(* Logix 5000 project; controller MV vendor 1 type 14 code 217 rev 31.11; software revision 31.00; part 29 of 53 *)
(* tags used below, declared in another part *)
   active : BOOL;
   Alarm_Reset : BOOL;
   CWD : CHECKWORD_FLAGS;
   Default_Check_Time : DINT;
   Item_Faults_Are_Latched : BOOL;
   Item_Simulation_Flag : BOOL;
   MC_CD_T2 : PlantItem;   // CD_T2
   MC_CH1_R1 : PlantItem;   // CH1_R1
   MC_CH1_R1_ALARM : ALARM_DIGITAL;
   MC_CH1_R1_C : ALIAS FOR RIO_Rack_2:4:I.Data.4;
   MC_CH1_R1_DR : ALIAS FOR RIO_Rack_2:5:O.Data.0;
   MC_CH1_R1_O : ALIAS FOR RIO_Rack_2:4:I.Data.0;
   MC_CH1_R1R : PlantItem;   // CH1_R1R
   MC_CH1_R1R_ALARM : ALARM_DIGITAL;
   MC_CH1_R1R_C : ALIAS FOR RIO_Rack_2:4:I.Data.14;
   MC_CH1_R1R_DR : ALIAS FOR RIO_Rack_2:5:O.Data.6;
   MC_CH1_R1R_O : ALIAS FOR RIO_Rack_2:4:I.Data.10;
   MC_CH1_R2 : PlantItem;   // CH1_R2
   MC_CH1_R2_ALARM : ALARM_DIGITAL;
   MC_CH1_R2_C : ALIAS FOR RIO_Rack_2:4:I.Data.5;
   MC_CH1_R2_DR : ALIAS FOR RIO_Rack_2:5:O.Data.1;
   MC_CH1_R2_O : ALIAS FOR RIO_Rack_2:4:I.Data.1;
   MC_CH1_R3 : PlantItem;   // CH1_R3
   MC_CH1_R3_ALARM : ALARM_DIGITAL;
   MC_CH1_R3_C : ALIAS FOR RIO_Rack_2:4:I.Data.6;
   MC_CH1_R3_DR : ALIAS FOR RIO_Rack_2:5:O.Data.2;
   MC_CH1_R3_O : ALIAS FOR RIO_Rack_2:4:I.Data.2;
   MC_CH1_R4 : PlantItem;   // CH1_R4
   MC_CH1_R4_ALARM : ALARM_DIGITAL;
   MC_CH1_R4_C : ALIAS FOR RIO_Rack_2:4:I.Data.7;
   MC_CH1_R4_DR : ALIAS FOR RIO_Rack_2:5:O.Data.3;
   MC_CH1_R4_O : ALIAS FOR RIO_Rack_2:4:I.Data.3;
   MC_CH1_R5 : PlantItem;   // CH1_R5
   MC_CH1_R5_ALARM : ALARM_DIGITAL;
   MC_CH1_R5_C : ALIAS FOR RIO_Rack_2:4:I.Data.12;
   MC_CH1_R5_DR : ALIAS FOR RIO_Rack_2:5:O.Data.4;
   MC_CH1_R5_O : ALIAS FOR RIO_Rack_2:4:I.Data.8;
   MC_CH1_R6 : PlantItem;   // CH1_R6
   MC_CH1_R6_ALARM : ALARM_DIGITAL;
   MC_CH1_R6_C : ALIAS FOR RIO_Rack_2:4:I.Data.13;
   MC_CH1_R6_DR : ALIAS FOR RIO_Rack_2:5:O.Data.5;
   MC_CH1_R6_O : ALIAS FOR RIO_Rack_2:4:I.Data.9;
   MC_FL_D2 : PlantItem;   // FL_D2
   MC_N10 : INT[255];   // SETTINGS
   MC_N100 : INT[255];   // C1_PLC Channel 1 PLC data
   MC_N104 : INT[255];   // CH1 REPORT Channel 1 CIP report file
   MC_N120 : INT[255];   // C2 PLC Channel 2 PLC data
   MC_N124 : INT[255];   // CH2 REPORT Channel 2 CIP report file
   MC_N200 : INT[255];   // CHK_WORK Plant item fault che cking work area
   MC_N7 : INT[255];   // INTEGER
   MC_N90 : INT[255];   // SV2_PLC Detergent tank 2 ser vice PLC data
   MC_N90_19_0_Storagebit : BOOL;
   MC_N90_32_0_Storagebit : BOOL;
   MC_N91 : INT[255];   // SV2_PC Detergent tank 2 ser vice PC to PLC data
   MC_P4 : PlantItem;   // P4
   MC_PROXY2 : PlantItem;   // PROXY2
   MC_SFile : INT[255];   // SLC Equivalent System File, So Original Code Can Remain
   MC_SV2 : PlantItem;   // SV2
   MC_T4 : TIMER[255];   // TIMER
   MC_T95 : TIMER[255];   // SV2 TIMERS
   One_Second_One_Scan : ALIAS FOR One_Second_1_scan;
(* MC_Common, continued *)

ROUTINE MC_SRV2_CMD_91   (* ladder *)
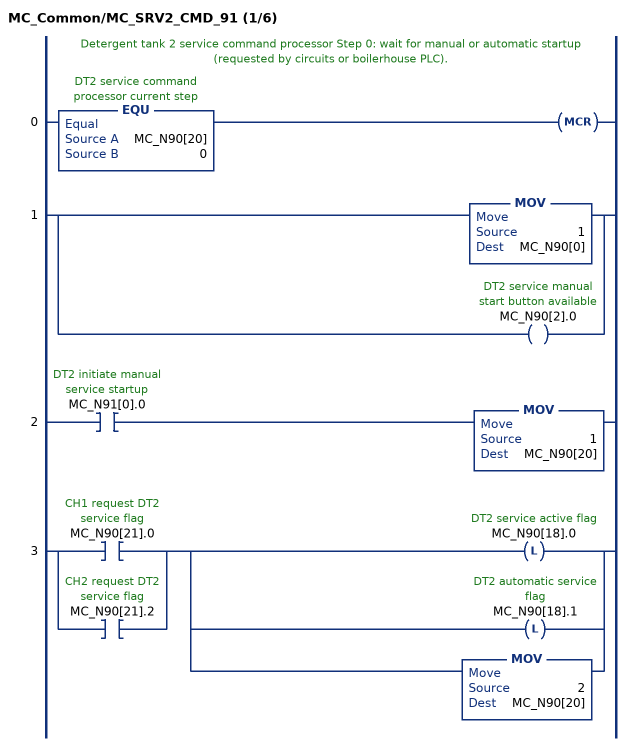
   // Detergent tank 2 service command processor Step 0: wait for manual or automatic startup (requested by circuits or boilerhouse PLC).
   0: EQU(MC_N90[20],0)MCR();
   1: [MOV(1,MC_N90[0]) ,OTE(MC_N90[2].0) ];
   2: XIC(MC_N91[0].0)MOV(1,MC_N90[20]);
   3: [XIC(MC_N90[21].0) ,XIC(MC_N90[21].2) ][OTL(MC_N90[18].0) ,OTL(MC_N90[18].1) ,MOV(2,MC_N90[20]) ];
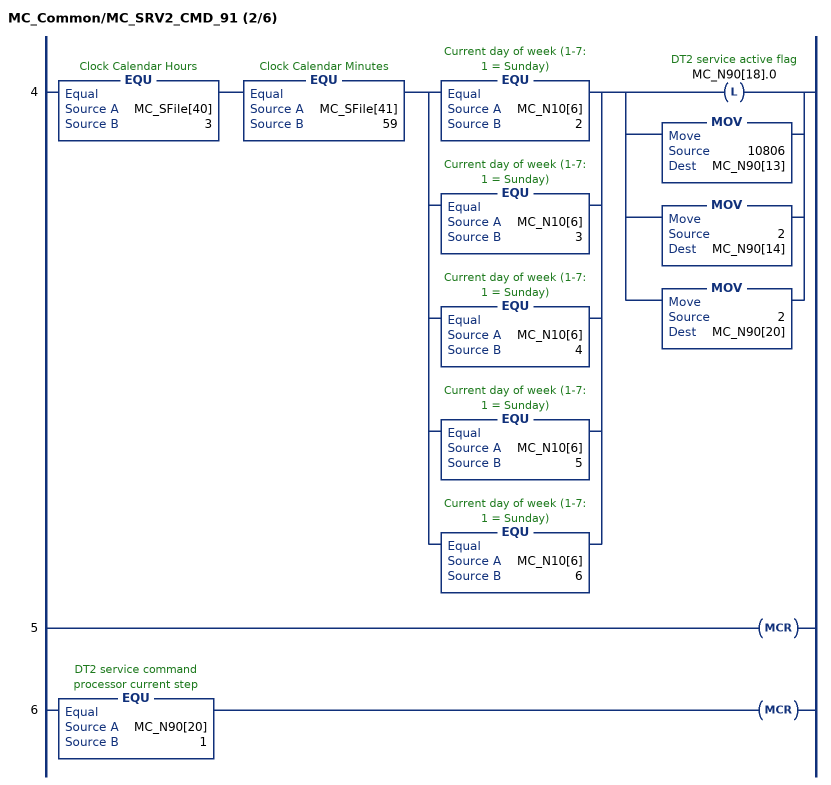
   4: EQU(MC_SFile[40],3)EQU(MC_SFile[41],59)[EQU(MC_N10[6],2) ,EQU(MC_N10[6],3) ,EQU(MC_N10[6],4) ,EQU(MC_N10[6],5) ,EQU(MC_N10[6],6) ][OTL(MC_N90[18].0) ,MOV(10806,MC_N90[13]) ,MOV(2,MC_N90[14]) ,MOV(2,MC_N90[20]) ];
   5: MCR();
   6: EQU(MC_N90[20],1)MCR();
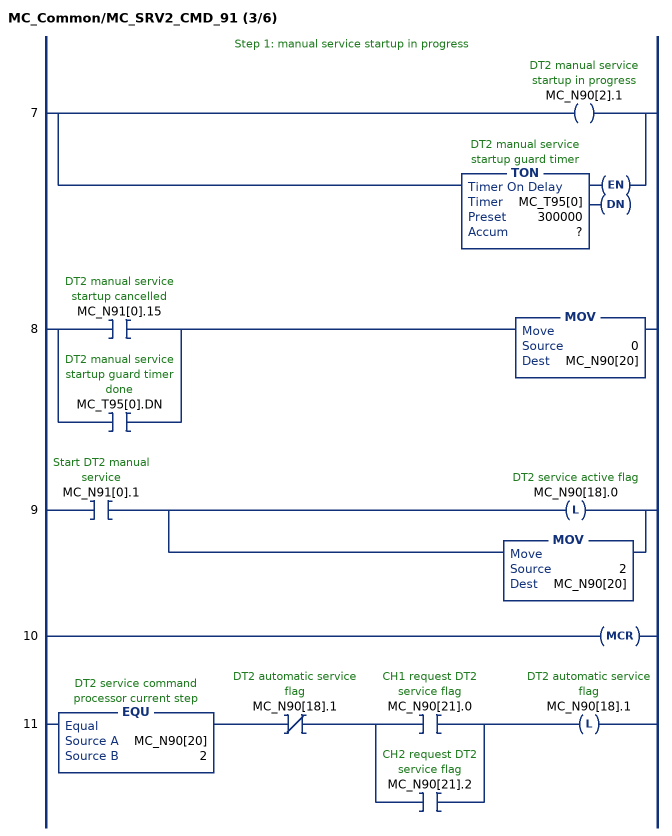
   // Step 1: manual service startup in progress
   7: [OTE(MC_N90[2].1) ,TON(MC_T95[0],?,?) ];
   8: [XIC(MC_N91[0].15) ,XIC(MC_T95[0].DN) ]MOV(0,MC_N90[20]);
   9: XIC(MC_N91[0].1)[OTL(MC_N90[18].0) ,MOV(2,MC_N90[20]) ];
   10: MCR();
   11: EQU(MC_N90[20],2)XIO(MC_N90[18].1)[XIC(MC_N90[21].0) ,XIC(MC_N90[21].2) ]OTL(MC_N90[18].1);
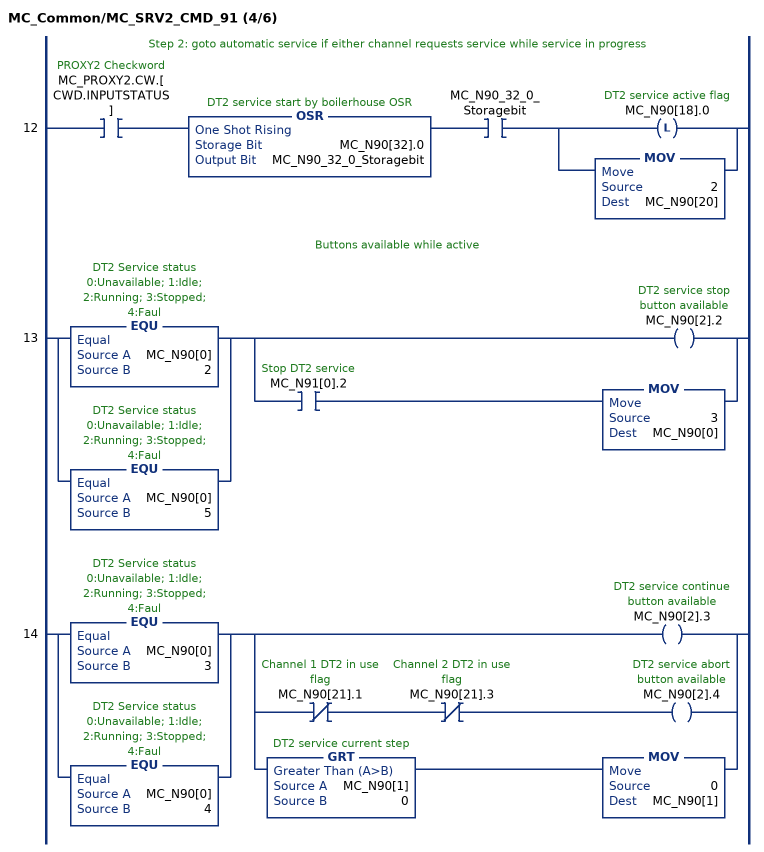
   // Step 2: goto automatic service if either channel requests service while service in progress
   12: XIC(MC_PROXY2.CW.[CWD.INPUTSTATUS])OSR(MC_N90[32].0,MC_N90_32_0_Storagebit)XIC(MC_N90_32_0_Storagebit)[OTL(MC_N90[18].0) ,MOV(2,MC_N90[20]) ];
   // Buttons available while active
   13: [EQU(MC_N90[0],2) ,EQU(MC_N90[0],5) ][OTE(MC_N90[2].2) ,XIC(MC_N91[0].2) MOV(3,MC_N90[0]) ];
   14: [EQU(MC_N90[0],3) ,EQU(MC_N90[0],4) ][OTE(MC_N90[2].3) ,XIO(MC_N90[21].1) XIO(MC_N90[21].3) OTE(MC_N90[2].4) ,GRT(MC_N90[1],0) MOV(0,MC_N90[1]) ];
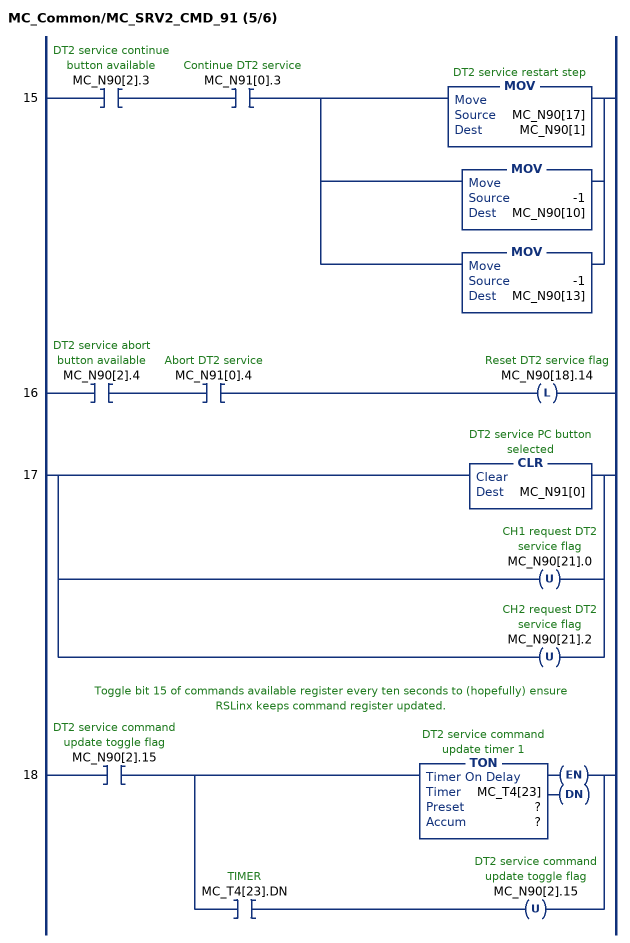
   15: XIC(MC_N90[2].3)XIC(MC_N91[0].3)[MOV(MC_N90[17],MC_N90[1]) ,MOV(-1,MC_N90[10]) ,MOV(-1,MC_N90[13]) ];
   16: XIC(MC_N90[2].4)XIC(MC_N91[0].4)OTL(MC_N90[18].14);
   17: [CLR(MC_N91[0]) ,OTU(MC_N90[21].0) ,OTU(MC_N90[21].2) ];
   // Toggle bit 15 of commands available register every ten seconds to (hopefully) ensure RSLinx keeps command register updated.
   18: XIC(MC_N90[2].15)[TON(MC_T4[23],?,?) ,XIC(MC_T4[23].DN) OTU(MC_N90[2].15) ];
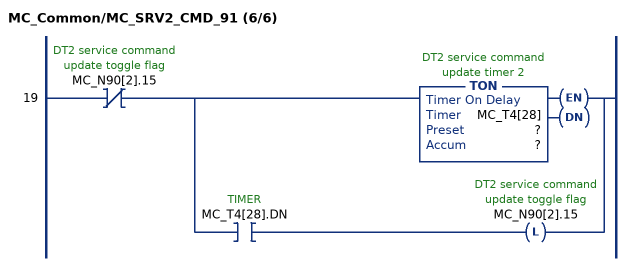
   19: XIO(MC_N90[2].15)[TON(MC_T4[28],?,?) ,XIC(MC_T4[28].DN) OTL(MC_N90[2].15) ];
END_ROUTINE

ROUTINE MC_SRV2_MCP_90   (* ladder *)
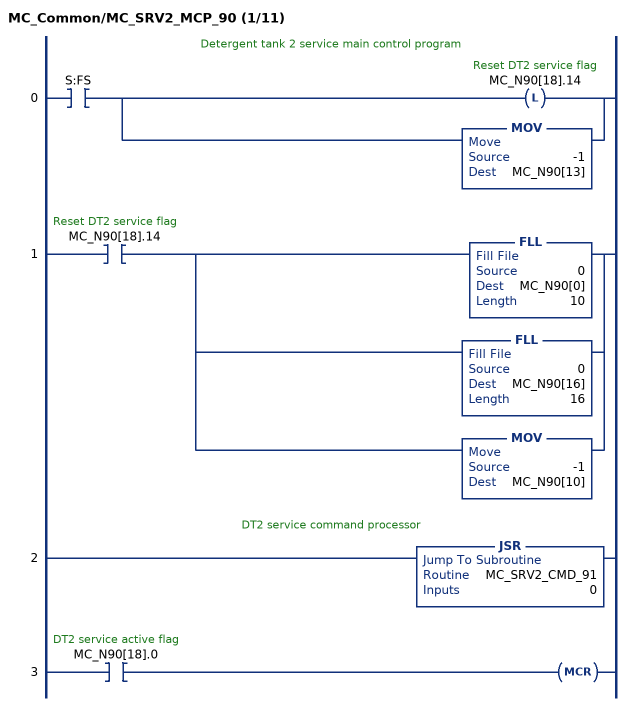
   // Detergent tank 2 service main control program
   0: XIC(S:FS)[OTL(MC_N90[18].14) ,MOV(-1,MC_N90[13]) ];
   1: XIC(MC_N90[18].14)[FLL(0,MC_N90[0],10) ,FLL(0,MC_N90[16],16) ,MOV(-1,MC_N90[10]) ];
   // DT2 service command processor
   2: JSR(MC_SRV2_CMD_91,0);
   3: XIC(MC_N90[18].0)MCR();
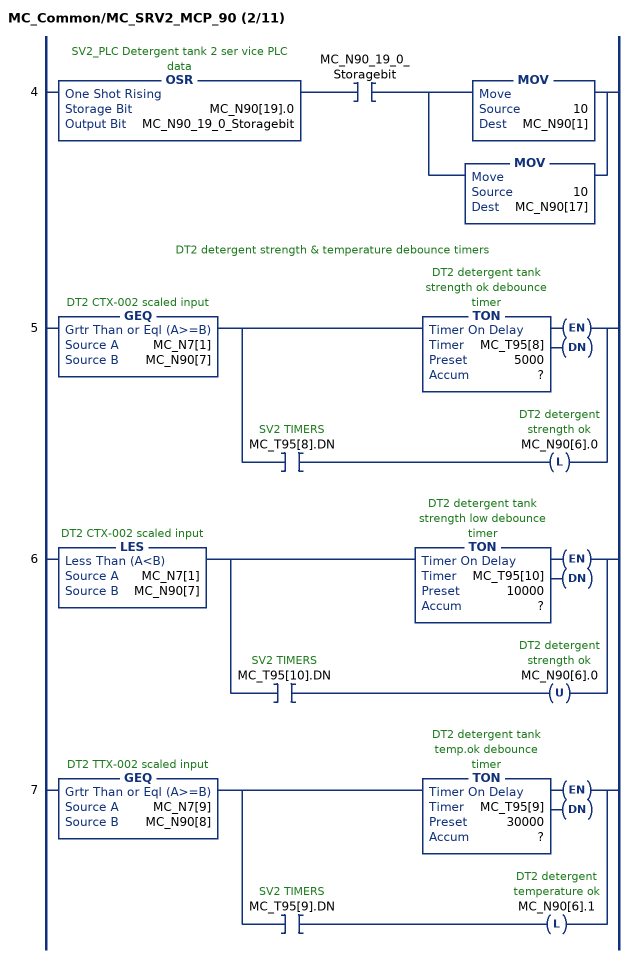
   4: OSR(MC_N90[19].0,MC_N90_19_0_Storagebit)XIC(MC_N90_19_0_Storagebit)[MOV(10,MC_N90[1]) ,MOV(10,MC_N90[17]) ];
   // DT2 detergent strength & temperature debounce timers
   5: GEQ(MC_N7[1],MC_N90[7])[TON(MC_T95[8],?,?) ,XIC(MC_T95[8].DN) OTL(MC_N90[6].0) ];
   6: LES(MC_N7[1],MC_N90[7])[TON(MC_T95[10],?,?) ,XIC(MC_T95[10].DN) OTU(MC_N90[6].0) ];
   7: GEQ(MC_N7[9],MC_N90[8])[TON(MC_T95[9],?,?) ,XIC(MC_T95[9].DN) OTL(MC_N90[6].1) ];
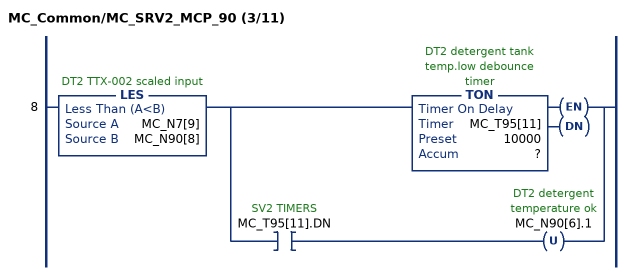
   8: LES(MC_N7[9],MC_N90[8])[TON(MC_T95[11],?,?) ,XIC(MC_T95[11].DN) OTU(MC_N90[6].1) ];
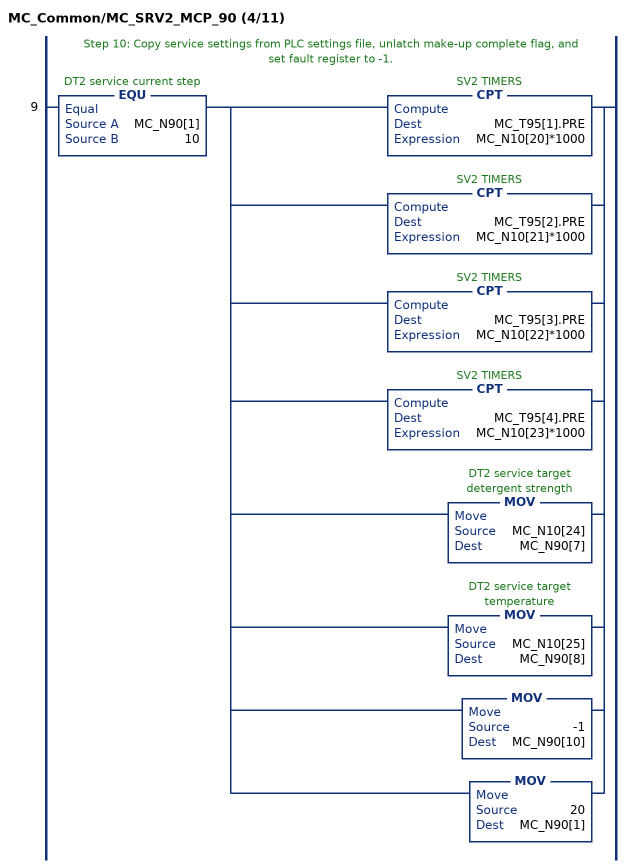
   // Step 10: Copy service settings from PLC settings file, unlatch make-up complete flag, and set fault register to -1.
   9: EQU(MC_N90[1],10)[CPT(MC_T95[1].PRE,MC_N10[20]*1000) ,CPT(MC_T95[2].PRE,MC_N10[21]*1000) ,CPT(MC_T95[3].PRE,MC_N10[22]*1000) ,CPT(MC_T95[4].PRE,MC_N10[23]*1000) ,MOV(MC_N10[24],MC_N90[7]) ,MOV(MC_N10[25],MC_N90[8]) ,MOV(-1,MC_N90[10]) ,MOV(20,MC_N90[1]) ];
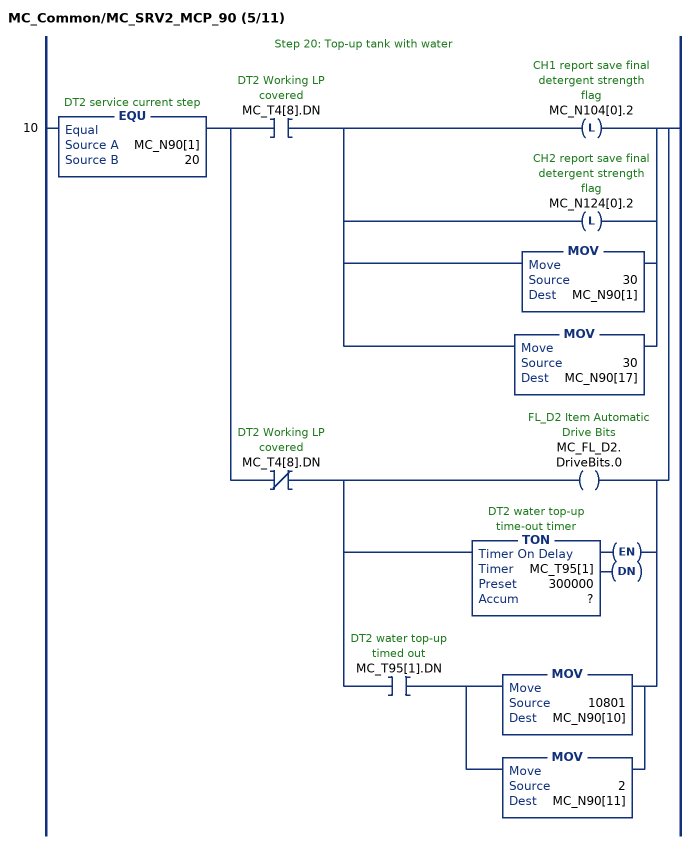
   // Step 20: Top-up tank with water
   10: EQU(MC_N90[1],20)[XIC(MC_T4[8].DN) [OTL(MC_N104[0].2) ,OTL(MC_N124[0].2) ,MOV(30,MC_N90[1]) ,MOV(30,MC_N90[17]) ] ,XIO(MC_T4[8].DN) [OTE(MC_FL_D2.DriveBits.0) ,TON(MC_T95[1],?,?) ,XIC(MC_T95[1].DN) [MOV(10801,MC_N90[10]) ,MOV(2,MC_N90[11]) ] ] ];
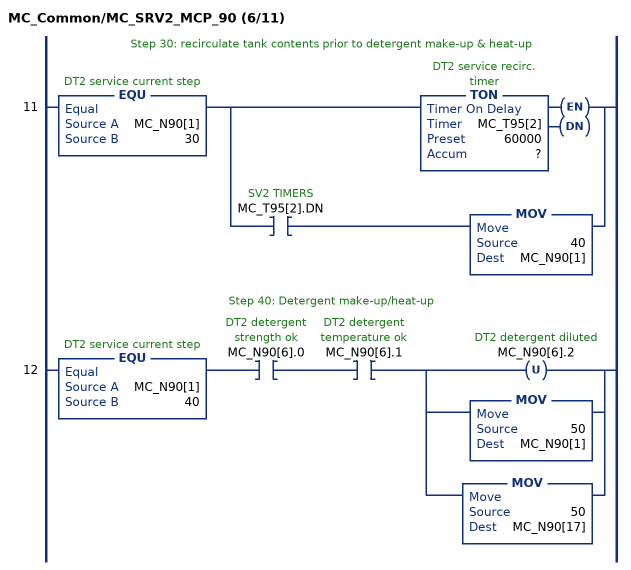
   // Step 30: recirculate tank contents prior to detergent make-up & heat-up
   11: EQU(MC_N90[1],30)[TON(MC_T95[2],?,?) ,XIC(MC_T95[2].DN) MOV(40,MC_N90[1]) ];
   // Step 40: Detergent make-up/heat-up
   12: EQU(MC_N90[1],40)XIC(MC_N90[6].0)XIC(MC_N90[6].1)[OTU(MC_N90[6].2) ,MOV(50,MC_N90[1]) ,MOV(50,MC_N90[17]) ];
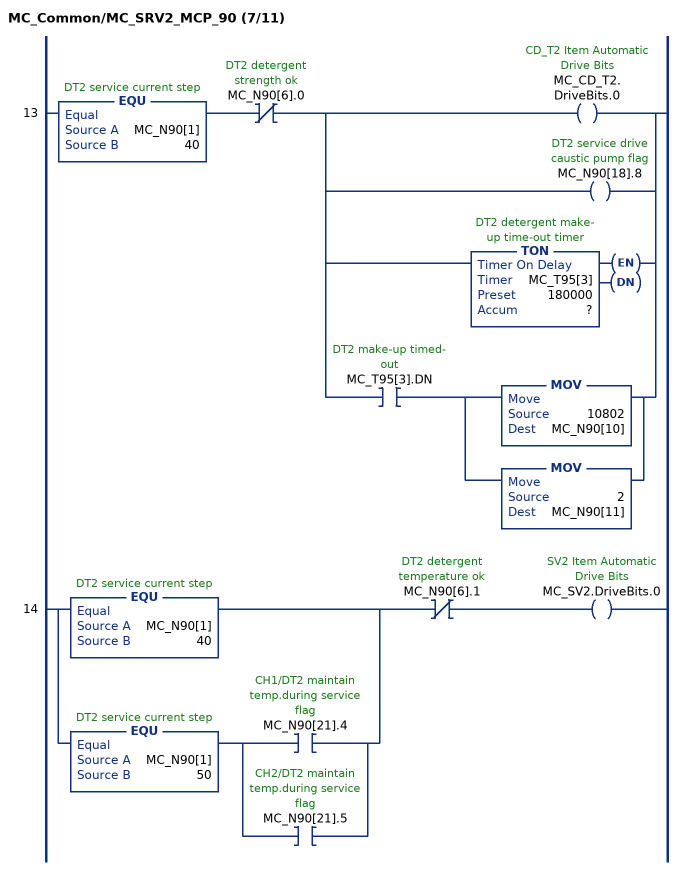
   13: EQU(MC_N90[1],40)XIO(MC_N90[6].0)[[OTE(MC_CD_T2.DriveBits.0) ,OTE(MC_N90[18].8) ] ,TON(MC_T95[3],?,?) ,XIC(MC_T95[3].DN) [MOV(10802,MC_N90[10]) ,MOV(2,MC_N90[11]) ] ];
   14: [EQU(MC_N90[1],40) ,EQU(MC_N90[1],50) [XIC(MC_N90[21].4) ,XIC(MC_N90[21].5) ] ]XIO(MC_N90[6].1)OTE(MC_SV2.DriveBits.0);
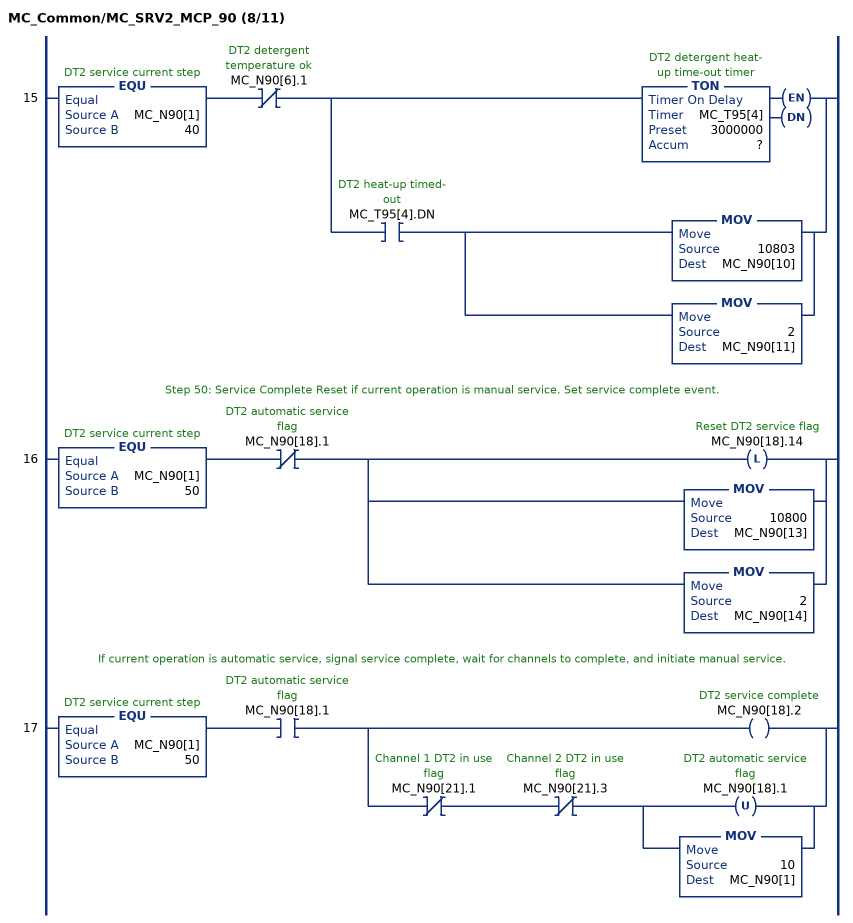
   15: EQU(MC_N90[1],40)XIO(MC_N90[6].1)[TON(MC_T95[4],?,?) ,XIC(MC_T95[4].DN) [MOV(10803,MC_N90[10]) ,MOV(2,MC_N90[11]) ] ];
   // Step 50: Service Complete Reset if current operation is manual service. Set service complete event.
   16: EQU(MC_N90[1],50)XIO(MC_N90[18].1)[OTL(MC_N90[18].14) ,MOV(10800,MC_N90[13]) ,MOV(2,MC_N90[14]) ];
   // If current operation is automatic service, signal service complete, wait for channels to complete, and initiate manual service.
   17: EQU(MC_N90[1],50)XIC(MC_N90[18].1)[OTE(MC_N90[18].2) ,XIO(MC_N90[21].1) XIO(MC_N90[21].3) [OTU(MC_N90[18].1) ,MOV(10,MC_N90[1]) ] ];
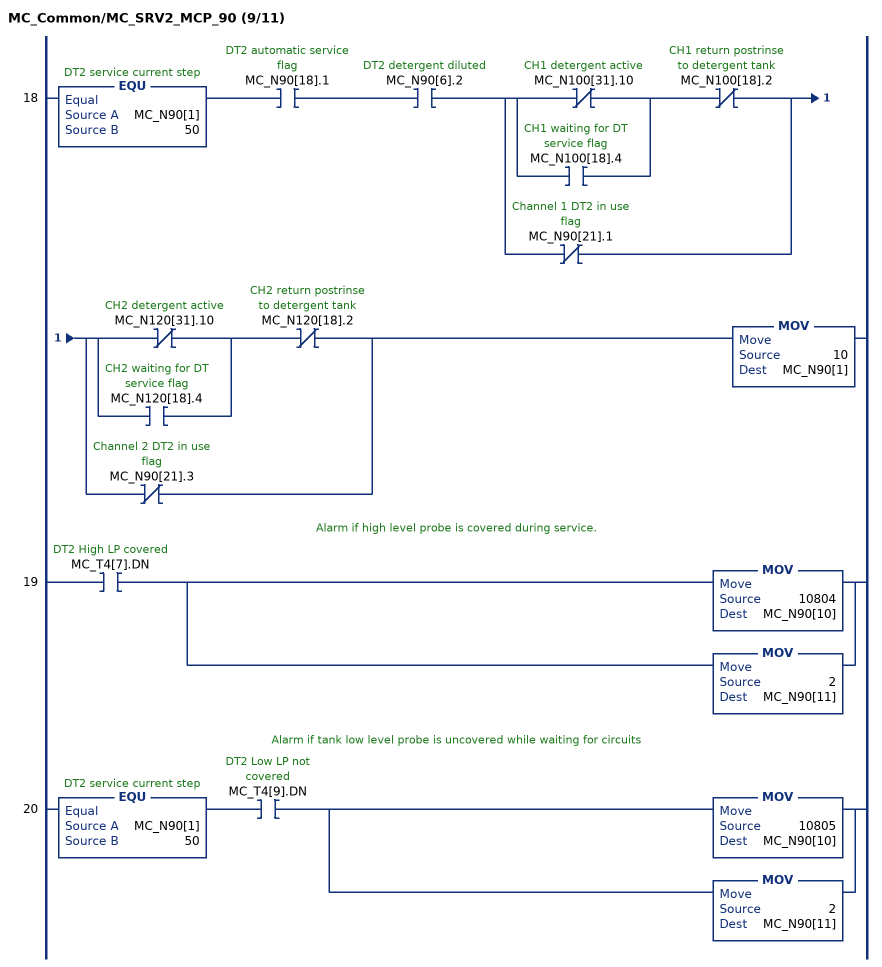
   18: EQU(MC_N90[1],50)XIC(MC_N90[18].1)XIC(MC_N90[6].2)[[XIO(MC_N100[31].10) ,XIC(MC_N100[18].4) ] XIO(MC_N100[18].2) ,XIO(MC_N90[21].1) ][[XIO(MC_N120[31].10) ,XIC(MC_N120[18].4) ] XIO(MC_N120[18].2) ,XIO(MC_N90[21].3) ]MOV(10,MC_N90[1]);
   // Alarm if high level probe is covered during service.
   19: XIC(MC_T4[7].DN)[MOV(10804,MC_N90[10]) ,MOV(2,MC_N90[11]) ];
   // Alarm if tank low level probe is uncovered while waiting for circuits
   20: EQU(MC_N90[1],50)XIC(MC_T4[9].DN)[MOV(10805,MC_N90[10]) ,MOV(2,MC_N90[11]) ];